        .Step_20   // Remove Lift comand
        .Step_03   // Rack Unlock Valve
        .Step_21   // Remove Unlock Comand
        .Step_04   // Lapbars Opening Valve -Y31008I
        .Step_22   // Lift comand
   RESTRAINTS_Left_Press_Switch_Series : BOOL := 1;
   RESTRAINTS_MainValve_PressTest : Valve_2_pos_monostable := (FeedBack_Type := 1, Discrepancy_Time := 2000, I_FeedBack_Data := 1, I_FeedBack_Status := 1, I_Output_Status := 1);
   RESTRAINTS_No_Alarms : BOOL := 1;
   RESTRAINTS_Open_Cycle_Ok : BOOL := 1;
   RESTRAINTS_Open_Postion : BOOL[64];
        [10]   // -B53201J
        [11]   // -B55001J
        [12]   // -B55007J
        [13]   // -B55101J
        [14]   // -B55107J
        [15]   // -B55201J
        [16]   // -B57001J
        [17]   // -B57007J
        [18]   // -B57101J
        [19]   // -B57107J
        [20]   // -B57201J
        [21]   // -B59001J
        [22]   // -B59007J
        [23]   // -B59101J
        [24]   // -B59107J
        [25]   // -B59201J
        [26]   // -B61001J
        [27]   // -B61007J
        [1]   // -B51001J
        [28]   // -B61101J
        [2]   // -B51007J
        [3]   // -B51101J
        [4]   // -B51107J
        [5]   // -B51201J
        [6]   // -B53001J
        [7]   // -B53007J
        [30]   // -B61201J
        [31]   // -B63001J
        [32]   // -B63007J
        [33]   // -B63101J
        [34]   // -B63107J
        [35]   // -B63201J
        [36]   // -B65001J
        [37]   // -B65007J
        [38]   // -B65101J
        [39]   // -B65007J
        [8]   // B53101J
        [9]   // B53107J
        [40]   // -B65201J
        [29]   // -B611017J
   RESTRAINTS_OpenComand : BOOL;   // Steps 01, 02, 03, 04
   RESTRAINTS_Opening : BOOL;
   Restraints_Permissive : Permissive := (All_Permissive_Ok := 1, BitsConditions := -1);
   Restraints_Permissive_Ok : BOOL := 1;
   Restraints_PermissiveLost : DINT := -2097153;
   RESTRAINTS_PressureSwitch_Working : BOOL := 1;
   RESTRAINTS_Rack : LapBar_Racks[41] := ([1].Input_Left.Discrepancy_Time := 3000, [1].Input_Left.Channel_A := 1, [1].Input_Left.Channel_B := 1, [1].Input_Left.Channel_A_Status := 1, [1].Input_Left.Channel_B_Status := 1, [1].Input_Left.O1 := 1, [1].Input_Right.Discrepancy_Time := 3000, [1].Input_Right.Channel_A := 1, [1].Input_Right.Channel_B := 1, [1].Input_Right.Channel_A_Status := 1, [1].Input_Right.Channel_B_Status := 1, [1].Input_Right.O1 := 1, [1].ON_Delay_Left.PRE := 500, [1].ON_Delay_Right.PRE := 500, [1].Memory_Left := 1, [1].Memory_Right := 1, [1].Memory_Left_Unlocked := 1, [1].Memory_Right_Unlocked := 1, [2].Input_Left.Discrepancy_Time := 3000, [2].Input_Left.Channel_A := 1, [2].Input_Left.Channel_B := 1, [2].Input_Left.Channel_A_Status := 1, [2].Input_Left.Channel_B_Status := 1, [2].Input_Left.O1 := 1, [2].Input_Right.Discrepancy_Time := 3000, [2].Input_Right.Channel_A := 1, [2].Input_Right.Channel_B := 1, [2].Input_Right.Channel_A_Status := 1, [2].Input_Right.Channel_B_Status := 1, [2].Input_Right.O1 := 1, [2].ON_Delay_Left.PRE := 500, [2].ON_Delay_Right.PRE := 500, [2].Memory_Left := 1, [2].Memory_Right := 1, [2].Memory_Left_Unlocked := 1, [2].Memory_Right_Unlocked := 1, [3].Input_Left.Discrepancy_Time := 3000, [3].Input_Left.Channel_A := 1, [3].Input_Left.Channel_B := 1, [3].Input_Left.Channel_A_Status := 1, [3].Input_Left.Channel_B_Status := 1, [3].Input_Left.O1 := 1, [3].Input_Right.Discrepancy_Time := 3000, [3].Input_Right.Channel_A := 1, [3].Input_Right.Channel_B := 1, [3].Input_Right.Channel_A_Status := 1, [3].Input_Right.Channel_B_Status := 1, [3].Input_Right.O1 := 1, [3].ON_Delay_Left.PRE := 500, [3].ON_Delay_Right.PRE := 500, [3].Memory_Left := 1, [3].Memory_Right := 1, [3].Memory_Left_Unlocked := 1, [3].Memory_Right_Unlocked := 1, [4].Input_Left.Discrepancy_Time := 3000, [4].Input_Left.Channel_A := 1, [4].Input_Left.Channel_B := 1, [4].Input_Left.Channel_A_Status := 1, [4].Input_Left.Channel_B_Status := 1, [4].Input_Left.O1 := 1,
        [4].Input_Right.Discrepancy_Time := 3000, [4].Input_Right.Channel_A := 1, [4].Input_Right.Channel_B := 1, [4].Input_Right.Channel_A_Status := 1, [4].Input_Right.Channel_B_Status := 1, [4].Input_Right.O1 := 1, [4].ON_Delay_Left.PRE := 500, [4].ON_Delay_Right.PRE := 500, [4].Memory_Left := 1, [4].Memory_Right := 1, [4].Memory_Left_Unlocked := 1, [4].Memory_Right_Unlocked := 1, [5].Input_Left.Discrepancy_Time := 3000, [5].Input_Left.Channel_A := 1, [5].Input_Left.Channel_B := 1, [5].Input_Left.Channel_A_Status := 1, [5].Input_Left.Channel_B_Status := 1, [5].Input_Left.O1 := 1, [5].Input_Right.Discrepancy_Time := 3000, [5].Input_Right.Channel_A := 1, [5].Input_Right.Channel_B := 1, [5].Input_Right.Channel_A_Status := 1, [5].Input_Right.Channel_B_Status := 1, [5].Input_Right.O1 := 1, [5].ON_Delay_Left.PRE := 500, [5].ON_Delay_Right.PRE := 500, [5].Memory_Left := 1, [5].Memory_Right := 1, [5].Memory_Left_Unlocked := 1, [5].Memory_Right_Unlocked := 1, [6].Input_Left.Discrepancy_Time := 3000, [6].Input_Left.Channel_A := 1, [6].Input_Left.Channel_B := 1, [6].Input_Left.Channel_A_Status := 1, [6].Input_Left.Channel_B_Status := 1, [6].Input_Left.O1 := 1, [6].Input_Right.Discrepancy_Time := 3000, [6].Input_Right.Channel_A := 1, [6].Input_Right.Channel_B := 1, [6].Input_Right.Channel_A_Status := 1, [6].Input_Right.Channel_B_Status := 1, [6].Input_Right.O1 := 1, [6].ON_Delay_Left.PRE := 500, [6].ON_Delay_Right.PRE := 500, [6].Memory_Left := 1, [6].Memory_Right := 1, [6].Memory_Left_Unlocked := 1, [6].Memory_Right_Unlocked := 1, [7].Input_Left.Discrepancy_Time := 3000, [7].Input_Left.Channel_A := 1, [7].Input_Left.Channel_B := 1, [7].Input_Left.Channel_A_Status := 1, [7].Input_Left.Channel_B_Status := 1, [7].Input_Left.O1 := 1, [7].Input_Right.Discrepancy_Time := 3000, [7].Input_Right.Channel_A := 1, [7].Input_Right.Channel_B := 1, [7].Input_Right.Channel_A_Status := 1, [7].Input_Right.Channel_B_Status := 1, [7].Input_Right.O1 := 1,
        [7].ON_Delay_Left.PRE := 500, [7].ON_Delay_Right.PRE := 500, [7].Memory_Left := 1, [7].Memory_Right := 1, [7].Memory_Left_Unlocked := 1, [7].Memory_Right_Unlocked := 1, [8].Input_Left.Discrepancy_Time := 3000, [8].Input_Left.Channel_A := 1, [8].Input_Left.Channel_B := 1, [8].Input_Left.Channel_A_Status := 1, [8].Input_Left.Channel_B_Status := 1, [8].Input_Left.O1 := 1, [8].Input_Right.Discrepancy_Time := 3000, [8].Input_Right.Channel_A := 1, [8].Input_Right.Channel_B := 1, [8].Input_Right.Channel_A_Status := 1, [8].Input_Right.Channel_B_Status := 1, [8].Input_Right.O1 := 1, [8].ON_Delay_Left.PRE := 500, [8].ON_Delay_Right.PRE := 500, [8].Memory_Left := 1, [8].Memory_Right := 1, [8].Memory_Left_Unlocked := 1, [8].Memory_Right_Unlocked := 1, [9].Input_Left.Discrepancy_Time := 3000, [9].Input_Left.Channel_A := 1, [9].Input_Left.Channel_B := 1, [9].Input_Left.Channel_A_Status := 1, [9].Input_Left.Channel_B_Status := 1, [9].Input_Left.O1 := 1, [9].Input_Right.Discrepancy_Time := 3000, [9].Input_Right.Channel_A_Status := 1, [9].Input_Right.Channel_B_Status := 1, [9].ON_Delay_Left.PRE := 500, [9].ON_Delay_Right.PRE := 500, [9].Memory_Left := 1, [9].Memory_Right := 1, [9].Memory_Left_Unlocked := 1, [9].Memory_Right_Unlocked := 1, [10].Input_Left.Discrepancy_Time := 3000, [10].Input_Left.Channel_A := 1, [10].Input_Left.Channel_B := 1, [10].Input_Left.Channel_A_Status := 1, [10].Input_Left.Channel_B_Status := 1, [10].Input_Left.O1 := 1, [10].Input_Right.Discrepancy_Time := 3000, [10].Input_Right.Channel_A := 1, [10].Input_Right.Channel_B := 1, [10].Input_Right.Channel_A_Status := 1, [10].Input_Right.Channel_B_Status := 1, [10].Input_Right.O1 := 1, [10].ON_Delay_Left.PRE := 500, [10].ON_Delay_Right.PRE := 500, [10].Memory_Left := 1, [10].Memory_Right := 1, [10].Memory_Left_Unlocked := 1, [10].Memory_Right_Unlocked := 1, [11].Input_Left.Discrepancy_Time := 3000, [11].Input_Left.Channel_A := 1, [11].Input_Left.Channel_B := 1,
        [11].Input_Left.Channel_A_Status := 1, [11].Input_Left.Channel_B_Status := 1, [11].Input_Left.O1 := 1, [11].Input_Right.Discrepancy_Time := 3000, [11].Input_Right.Channel_A := 1, [11].Input_Right.Channel_B := 1, [11].Input_Right.Channel_A_Status := 1, [11].Input_Right.Channel_B_Status := 1, [11].Input_Right.O1 := 1, [11].ON_Delay_Left.PRE := 500, [11].ON_Delay_Right.PRE := 500, [11].Memory_Left := 1, [11].Memory_Right := 1, [11].Memory_Left_Unlocked := 1, [11].Memory_Right_Unlocked := 1, [12].Input_Left.Discrepancy_Time := 3000, [12].Input_Left.Channel_A := 1, [12].Input_Left.Channel_B := 1, [12].Input_Left.Channel_A_Status := 1, [12].Input_Left.Channel_B_Status := 1, [12].Input_Left.O1 := 1, [12].Input_Right.Discrepancy_Time := 3000, [12].Input_Right.Channel_A := 1, [12].Input_Right.Channel_B := 1, [12].Input_Right.Channel_A_Status := 1, [12].Input_Right.Channel_B_Status := 1, [12].Input_Right.O1 := 1, [12].ON_Delay_Left.PRE := 500, [12].ON_Delay_Right.PRE := 500, [12].Memory_Left := 1, [12].Memory_Right := 1, [12].Memory_Left_Unlocked := 1, [12].Memory_Right_Unlocked := 1, [13].Input_Left.Discrepancy_Time := 3000, [13].Input_Left.Channel_A := 1, [13].Input_Left.Channel_B := 1, [13].Input_Left.Channel_A_Status := 1, [13].Input_Left.Channel_B_Status := 1, [13].Input_Left.O1 := 1, [13].Input_Right.Discrepancy_Time := 3000, [13].Input_Right.Channel_A := 1, [13].Input_Right.Channel_B := 1, [13].Input_Right.Channel_A_Status := 1, [13].Input_Right.Channel_B_Status := 1, [13].Input_Right.O1 := 1, [13].ON_Delay_Left.PRE := 500, [13].ON_Delay_Right.PRE := 500, [13].Memory_Left := 1, [13].Memory_Right := 1, [13].Memory_Left_Unlocked := 1, [13].Memory_Right_Unlocked := 1, [14].Input_Left.Discrepancy_Time := 3000, [14].Input_Left.Channel_A := 1, [14].Input_Left.Channel_B := 1, [14].Input_Left.Channel_A_Status := 1, [14].Input_Left.Channel_B_Status := 1, [14].Input_Left.O1 := 1, [14].Input_Right.Discrepancy_Time := 3000, [14].Input_Right.Channel_A := 1, [14].Input_Right.Channel_B := 1,
        [14].Input_Right.Channel_A_Status := 1, [14].Input_Right.Channel_B_Status := 1, [14].Input_Right.O1 := 1, [14].ON_Delay_Left.PRE := 500, [14].ON_Delay_Right.PRE := 500, [14].Memory_Left := 1, [14].Memory_Right := 1, [14].Memory_Left_Unlocked := 1, [14].Memory_Right_Unlocked := 1, [15].Input_Left.Discrepancy_Time := 3000, [15].Input_Left.Channel_A := 1, [15].Input_Left.Channel_B := 1, [15].Input_Left.Channel_A_Status := 1, [15].Input_Left.Channel_B_Status := 1, [15].Input_Left.O1 := 1, [15].Input_Right.Discrepancy_Time := 3000, [15].Input_Right.Channel_A := 1, [15].Input_Right.Channel_B := 1, [15].Input_Right.Channel_A_Status := 1, [15].Input_Right.Channel_B_Status := 1, [15].Input_Right.O1 := 1, [15].ON_Delay_Left.PRE := 500, [15].ON_Delay_Right.PRE := 500, [15].Memory_Left := 1, [15].Memory_Right := 1, [15].Memory_Left_Unlocked := 1, [15].Memory_Right_Unlocked := 1, [16].Input_Left.Discrepancy_Time := 3000, [16].Input_Left.Channel_A := 1, [16].Input_Left.Channel_B := 1, [16].Input_Left.Channel_A_Status := 1, [16].Input_Left.Channel_B_Status := 1, [16].Input_Left.O1 := 1, [16].Input_Right.Discrepancy_Time := 3000, [16].Input_Right.Channel_A := 1, [16].Input_Right.Channel_B := 1, [16].Input_Right.Channel_A_Status := 1, [16].Input_Right.Channel_B_Status := 1, [16].Input_Right.O1 := 1, [16].ON_Delay_Left.PRE := 500, [16].ON_Delay_Right.PRE := 500, [16].Memory_Left := 1, [16].Memory_Right := 1, [16].Memory_Left_Unlocked := 1, [16].Memory_Right_Unlocked := 1, [17].Input_Left.Discrepancy_Time := 3000, [17].Input_Left.Channel_A := 1, [17].Input_Left.Channel_B := 1, [17].Input_Left.Channel_A_Status := 1, [17].Input_Left.Channel_B_Status := 1, [17].Input_Left.O1 := 1, [17].Input_Right.Discrepancy_Time := 3000, [17].Input_Right.Channel_A := 1, [17].Input_Right.Channel_B := 1, [17].Input_Right.Channel_A_Status := 1, [17].Input_Right.Channel_B_Status := 1, [17].Input_Right.O1 := 1, [17].ON_Delay_Left.PRE := 500, [17].ON_Delay_Right.PRE := 500, [17].Memory_Left := 1,
        [17].Memory_Right := 1, [18].Input_Left.Discrepancy_Time := 3000, [18].Input_Left.Channel_A := 1, [18].Input_Left.Channel_B := 1, [18].Input_Left.Channel_A_Status := 1, [18].Input_Left.Channel_B_Status := 1, [18].Input_Left.O1 := 1, [18].Input_Right.Discrepancy_Time := 3000, [18].Input_Right.Channel_A := 1, [18].Input_Right.Channel_B := 1, [18].Input_Right.Channel_A_Status := 1, [18].Input_Right.Channel_B_Status := 1, [18].Input_Right.O1 := 1, [18].ON_Delay_Left.PRE := 500, [18].ON_Delay_Right.PRE := 500, [18].Memory_Left := 1, [18].Memory_Right := 1, [19].Input_Left.Discrepancy_Time := 3000, [19].Input_Left.Channel_A := 1, [19].Input_Left.Channel_B := 1, [19].Input_Left.Channel_A_Status := 1, [19].Input_Left.Channel_B_Status := 1, [19].Input_Left.O1 := 1, [19].Input_Right.Discrepancy_Time := 3000, [19].Input_Right.Channel_A := 1, [19].Input_Right.Channel_B := 1, [19].Input_Right.Channel_A_Status := 1, [19].Input_Right.Channel_B_Status := 1, [19].Input_Right.O1 := 1, [19].ON_Delay_Left.PRE := 500, [19].ON_Delay_Right.PRE := 500, [19].Memory_Left := 1, [19].Memory_Right := 1, [20].Input_Left.Discrepancy_Time := 3000, [20].Input_Left.Channel_A := 1, [20].Input_Left.Channel_B := 1, [20].Input_Left.Channel_A_Status := 1, [20].Input_Left.Channel_B_Status := 1, [20].Input_Left.O1 := 1, [20].Input_Right.Discrepancy_Time := 3000, [20].Input_Right.Channel_A := 1, [20].Input_Right.Channel_B := 1, [20].Input_Right.Channel_A_Status := 1, [20].Input_Right.Channel_B_Status := 1, [20].Input_Right.O1 := 1, [20].ON_Delay_Left.PRE := 500, [20].ON_Delay_Right.PRE := 500, [20].Memory_Left := 1, [20].Memory_Right := 1, [21].Input_Left.Discrepancy_Time := 3000, [21].Input_Left.Channel_A := 1, [21].Input_Left.Channel_B := 1, [21].Input_Left.Channel_A_Status := 1, [21].Input_Left.Channel_B_Status := 1, [21].Input_Left.O1 := 1, [21].Input_Right.Discrepancy_Time := 3000, [21].Input_Right.Channel_A := 1, [21].Input_Right.Channel_B := 1, [21].Input_Right.Channel_A_Status := 1, [21].Input_Right.Channel_B_Status := 1,
        [21].Input_Right.O1 := 1, [21].ON_Delay_Left.PRE := 500, [21].ON_Delay_Right.PRE := 500, [21].Memory_Left := 1, [21].Memory_Right := 1, [22].Input_Left.Discrepancy_Time := 3000, [22].Input_Left.Channel_A := 1, [22].Input_Left.Channel_B := 1, [22].Input_Left.Channel_A_Status := 1, [22].Input_Left.Channel_B_Status := 1, [22].Input_Left.O1 := 1, [22].Input_Right.Discrepancy_Time := 3000, [22].Input_Right.Channel_A := 1, [22].Input_Right.Channel_B := 1, [22].Input_Right.Channel_A_Status := 1, [22].Input_Right.Channel_B_Status := 1, [22].Input_Right.O1 := 1, [22].ON_Delay_Left.PRE := 500, [22].ON_Delay_Right.PRE := 500, [22].Memory_Left := 1, [22].Memory_Right := 1, [23].Input_Left.Discrepancy_Time := 3000, [23].Input_Left.Channel_A := 1, [23].Input_Left.Channel_B := 1, [23].Input_Left.Channel_A_Status := 1, [23].Input_Left.Channel_B_Status := 1, [23].Input_Left.O1 := 1, [23].Input_Right.Discrepancy_Time := 3000, [23].Input_Right.Channel_A := 1, [23].Input_Right.Channel_B := 1, [23].Input_Right.Channel_A_Status := 1, [23].Input_Right.Channel_B_Status := 1, [23].Input_Right.O1 := 1, [23].ON_Delay_Left.PRE := 500, [23].ON_Delay_Right.PRE := 500, [23].Memory_Left := 1, [23].Memory_Right := 1, [24].Input_Left.Discrepancy_Time := 3000, [24].Input_Left.Channel_A := 1, [24].Input_Left.Channel_B := 1, [24].Input_Left.Channel_A_Status := 1, [24].Input_Left.Channel_B_Status := 1, [24].Input_Left.O1 := 1, [24].Input_Right.Discrepancy_Time := 3000, [24].Input_Right.Channel_A := 1, [24].Input_Right.Channel_B := 1, [24].Input_Right.Channel_A_Status := 1, [24].Input_Right.Channel_B_Status := 1, [24].Input_Right.O1 := 1, [24].ON_Delay_Left.PRE := 500, [24].ON_Delay_Right.PRE := 500, [24].Memory_Left := 1, [24].Memory_Right := 1, [25].Input_Left.Discrepancy_Time := 3000, [25].Input_Left.Channel_A := 1, [25].Input_Left.Channel_B := 1, [25].Input_Left.Channel_A_Status := 1, [25].Input_Left.Channel_B_Status := 1, [25].Input_Left.O1 := 1, [25].Input_Right.Discrepancy_Time := 3000,
        [25].Input_Right.Channel_A := 1, [25].Input_Right.Channel_B := 1, [25].Input_Right.Channel_A_Status := 1, [25].Input_Right.Channel_B_Status := 1, [25].Input_Right.O1 := 1, [25].ON_Delay_Left.PRE := 500, [25].ON_Delay_Right.PRE := 500, [25].Memory_Left := 1, [25].Memory_Right := 1, [26].Input_Left.Discrepancy_Time := 3000, [26].Input_Left.Channel_A := 1, [26].Input_Left.Channel_B := 1, [26].Input_Left.Channel_A_Status := 1, [26].Input_Left.Channel_B_Status := 1, [26].Input_Left.O1 := 1, [26].Input_Right.Discrepancy_Time := 3000, [26].Input_Right.Channel_A := 1, [26].Input_Right.Channel_B := 1, [26].Input_Right.Channel_A_Status := 1, [26].Input_Right.Channel_B_Status := 1, [26].Input_Right.O1 := 1, [26].ON_Delay_Left.PRE := 500, [26].ON_Delay_Right.PRE := 500, [26].Memory_Left := 1, [26].Memory_Right := 1, [27].Input_Left.Discrepancy_Time := 3000, [27].Input_Left.Channel_A := 1, [27].Input_Left.Channel_B := 1, [27].Input_Left.Channel_A_Status := 1, [27].Input_Left.Channel_B_Status := 1, [27].Input_Left.O1 := 1, [27].Input_Right.Discrepancy_Time := 3000, [27].Input_Right.Channel_A := 1, [27].Input_Right.Channel_B := 1, [27].Input_Right.Channel_A_Status := 1, [27].Input_Right.Channel_B_Status := 1, [27].Input_Right.O1 := 1, [27].ON_Delay_Left.PRE := 500, [27].ON_Delay_Right.PRE := 500, [27].Memory_Left := 1, [27].Memory_Right := 1, [28].Input_Left.Discrepancy_Time := 3000, [28].Input_Left.Channel_A := 1, [28].Input_Left.Channel_B := 1, [28].Input_Left.Channel_A_Status := 1, [28].Input_Left.Channel_B_Status := 1, [28].Input_Left.O1 := 1, [28].Input_Right.Discrepancy_Time := 3000, [28].Input_Right.Channel_A := 1, [28].Input_Right.Channel_B := 1, [28].Input_Right.Channel_A_Status := 1, [28].Input_Right.Channel_B_Status := 1, [28].Input_Right.O1 := 1, [28].ON_Delay_Left.PRE := 500, [28].ON_Delay_Right.PRE := 500, [28].Memory_Left := 1, [28].Memory_Right := 1, [29].Input_Left.Discrepancy_Time := 3000, [29].Input_Left.Channel_A := 1, [29].Input_Left.Channel_B := 1,
        [29].Input_Left.Channel_A_Status := 1, [29].Input_Left.Channel_B_Status := 1, [29].Input_Left.O1 := 1, [29].Input_Right.Discrepancy_Time := 3000, [29].Input_Right.Channel_A := 1, [29].Input_Right.Channel_B := 1, [29].Input_Right.Channel_A_Status := 1, [29].Input_Right.Channel_B_Status := 1, [29].Input_Right.O1 := 1, [29].ON_Delay_Left.PRE := 500, [29].ON_Delay_Right.PRE := 500, [29].Memory_Left := 1, [29].Memory_Right := 1, [30].Input_Left.Discrepancy_Time := 3000, [30].Input_Left.Channel_A := 1, [30].Input_Left.Channel_B := 1, [30].Input_Left.Channel_A_Status := 1, [30].Input_Left.Channel_B_Status := 1, [30].Input_Left.O1 := 1, [30].Input_Right.Discrepancy_Time := 3000, [30].Input_Right.Channel_A := 1, [30].Input_Right.Channel_B := 1, [30].Input_Right.Channel_A_Status := 1, [30].Input_Right.Channel_B_Status := 1, [30].Input_Right.O1 := 1, [30].ON_Delay_Left.PRE := 500, [30].ON_Delay_Right.PRE := 500, [30].Memory_Left := 1, [30].Memory_Right := 1, [31].Input_Left.Discrepancy_Time := 3000, [31].Input_Left.Channel_A := 1, [31].Input_Left.Channel_B := 1, [31].Input_Left.Channel_A_Status := 1, [31].Input_Left.Channel_B_Status := 1, [31].Input_Left.O1 := 1, [31].Input_Right.Discrepancy_Time := 3000, [31].Input_Right.Channel_A := 1, [31].Input_Right.Channel_B := 1, [31].Input_Right.Channel_A_Status := 1, [31].Input_Right.Channel_B_Status := 1, [31].Input_Right.O1 := 1, [31].ON_Delay_Left.PRE := 500, [31].ON_Delay_Right.PRE := 500, [31].Memory_Left := 1, [31].Memory_Right := 1, [32].Input_Left.Discrepancy_Time := 3000, [32].Input_Left.Channel_A := 1, [32].Input_Left.Channel_B := 1, [32].Input_Left.Channel_A_Status := 1, [32].Input_Left.Channel_B_Status := 1, [32].Input_Left.O1 := 1, [32].Input_Right.Discrepancy_Time := 3000, [32].Input_Right.Channel_A := 1, [32].Input_Right.Channel_B := 1, [32].Input_Right.Channel_A_Status := 1, [32].Input_Right.Channel_B_Status := 1, [32].Input_Right.O1 := 1, [32].ON_Delay_Left.PRE := 500, [32].ON_Delay_Right.PRE := 500, [32].Memory_Left := 1,
        [32].Memory_Right := 1, [33].Input_Left.Discrepancy_Time := 3000, [33].Input_Left.Channel_A := 1, [33].Input_Left.Channel_B := 1, [33].Input_Left.Channel_A_Status := 1, [33].Input_Left.Channel_B_Status := 1, [33].Input_Left.O1 := 1, [33].Input_Right.Discrepancy_Time := 3000, [33].Input_Right.Channel_A := 1, [33].Input_Right.Channel_B := 1, [33].Input_Right.Channel_A_Status := 1, [33].Input_Right.Channel_B_Status := 1, [33].Input_Right.O1 := 1, [33].ON_Delay_Left.PRE := 500, [33].ON_Delay_Right.PRE := 500, [33].Memory_Left := 1, [33].Memory_Right := 1, [34].Input_Left.Discrepancy_Time := 3000, [34].Input_Left.Channel_A := 1, [34].Input_Left.Channel_B := 1, [34].Input_Left.Channel_A_Status := 1, [34].Input_Left.Channel_B_Status := 1, [34].Input_Left.O1 := 1, [34].Input_Right.Discrepancy_Time := 3000, [34].Input_Right.Channel_A := 1, [34].Input_Right.Channel_B := 1, [34].Input_Right.Channel_A_Status := 1, [34].Input_Right.Channel_B_Status := 1, [34].Input_Right.O1 := 1, [34].ON_Delay_Left.PRE := 500, [34].ON_Delay_Right.PRE := 500, [34].Memory_Left := 1, [34].Memory_Right := 1, [35].Input_Left.Discrepancy_Time := 3000, [35].Input_Left.Channel_A := 1, [35].Input_Left.Channel_B := 1, [35].Input_Left.Channel_A_Status := 1, [35].Input_Left.Channel_B_Status := 1, [35].Input_Left.O1 := 1, [35].Input_Right.Discrepancy_Time := 3000, [35].Input_Right.Channel_A := 1, [35].Input_Right.Channel_B := 1, [35].Input_Right.Channel_A_Status := 1, [35].Input_Right.Channel_B_Status := 1, [35].Input_Right.O1 := 1, [35].ON_Delay_Left.PRE := 500, [35].ON_Delay_Right.PRE := 500, [35].Memory_Left := 1, [35].Memory_Right := 1, [36].Input_Left.Discrepancy_Time := 3000, [36].Input_Left.Channel_A := 1, [36].Input_Left.Channel_B := 1, [36].Input_Left.Channel_A_Status := 1, [36].Input_Left.Channel_B_Status := 1, [36].Input_Left.O1 := 1, [36].Input_Right.Discrepancy_Time := 3000, [36].Input_Right.Channel_A := 1, [36].Input_Right.Channel_B := 1, [36].Input_Right.Channel_A_Status := 1, [36].Input_Right.Channel_B_Status := 1,
        [36].Input_Right.O1 := 1, [36].ON_Delay_Left.PRE := 500, [36].ON_Delay_Right.PRE := 500, [36].Memory_Left := 1, [36].Memory_Right := 1, [37].Input_Left.Discrepancy_Time := 3000, [37].Input_Left.Channel_A := 1, [37].Input_Left.Channel_B := 1, [37].Input_Left.Channel_A_Status := 1, [37].Input_Left.Channel_B_Status := 1, [37].Input_Left.O1 := 1, [37].Input_Right.Discrepancy_Time := 3000, [37].Input_Right.Channel_A := 1, [37].Input_Right.Channel_B := 1, [37].Input_Right.Channel_A_Status := 1, [37].Input_Right.Channel_B_Status := 1, [37].Input_Right.O1 := 1, [37].ON_Delay_Left.PRE := 500, [37].ON_Delay_Right.PRE := 500, [37].Memory_Left := 1, [37].Memory_Right := 1, [38].Input_Left.Discrepancy_Time := 3000, [38].Input_Left.Channel_A := 1, [38].Input_Left.Channel_B := 1, [38].Input_Left.Channel_A_Status := 1, [38].Input_Left.Channel_B_Status := 1, [38].Input_Left.O1 := 1, [38].Input_Right.Discrepancy_Time := 3000, [38].Input_Right.Channel_A := 1, [38].Input_Right.Channel_B := 1, [38].Input_Right.Channel_A_Status := 1, [38].Input_Right.Channel_B_Status := 1, [38].Input_Right.O1 := 1, [38].ON_Delay_Left.PRE := 500, [38].ON_Delay_Right.PRE := 500, [38].Memory_Left := 1, [38].Memory_Right := 1, [39].Input_Left.Discrepancy_Time := 3000, [39].Input_Left.Channel_A := 1, [39].Input_Left.Channel_B := 1, [39].Input_Left.Channel_A_Status := 1, [39].Input_Left.Channel_B_Status := 1, [39].Input_Left.O1 := 1, [39].Input_Right.Discrepancy_Time := 3000, [39].Input_Right.Channel_A := 1, [39].Input_Right.Channel_B := 1, [39].Input_Right.Channel_A_Status := 1, [39].Input_Right.Channel_B_Status := 1, [39].Input_Right.O1 := 1, [39].ON_Delay_Left.PRE := 500, [39].ON_Delay_Right.PRE := 500, [39].Memory_Left := 1, [39].Memory_Right := 1, [40].Input_Left.Discrepancy_Time := 3000, [40].Input_Left.Channel_A := 1, [40].Input_Left.Channel_B := 1, [40].Input_Left.Channel_A_Status := 1, [40].Input_Left.Channel_B_Status := 1, [40].Input_Left.O1 := 1, [40].Input_Right.Discrepancy_Time := 3000,
        [40].Input_Right.Channel_A := 1, [40].Input_Right.Channel_B := 1, [40].Input_Right.Channel_A_Status := 1, [40].Input_Right.Channel_B_Status := 1, [40].Input_Right.O1 := 1, [40].ON_Delay_Left.PRE := 500, [40].ON_Delay_Right.PRE := 500, [40].Memory_Left := 1, [40].Memory_Right := 1);
        [10].Input_Left   // -A53702I
        [1].Input_Left   // -A51302I
        [10].Input_Right   // -A53707I
        [1].Input_Right   // -A51307I
        [2].Input_Left   // -A51402I
        [11].Input_Left   // -A55302I
        [2].Input_Right   // -A51407I
        [11].Input_Right   // -A55307I
        [12].Input_Left   // -A55402I
        [12].Input_Right   // -A55407I
        [13].Input_Left   // -A55502I
        [3].Input_Left   // -A51502I
        [13].Input_Right   // -A55507I
        [3].Input_Right   // -A51507I
        [4].Input_Left   // -A51602I
        [4].Input_Right   // -A51607I
        [5].Input_Left   // -A51702I
        [5].Input_Right   // -A51707I
        [6].Input_Left   // -A53302I
        [6].Input_Right   // -A53307I
        [7].Input_Left   // -A53402I
        [14].Input_Left   // -A55602I
        [7].Input_Right   // -A534027I
        [14].Input_Right   // -A55607I
        [15].Input_Left   // -A55702I
        [15].Input_Right   // -A55707I
        [8].Input_Left   // -A53502I
        [8].Input_Right   // -A53507I
        [9].Input_Left   // -A53602I
        [9].Input_Right   // -A53607I
        [16].Input_Left   // -A57402I
        [16].Input_Right   // -A57407I
        [17].Input_Left   // -A57402I
        [17].Input_Right   // -A57407I
        [18].Input_Left   // -A57502I
        [18].Input_Right   // -A57507I
        [19].Input_Left   // -A57602I
        [19].Input_Right   // -A57607I
        [20].Input_Left   // -A57702I
        [20].Input_Right   // -A57707I
        [21].Input_Left   // -A59302I
        [21].Input_Right   // -A59307I
        [22].Input_Left   // -A59402I
        [22].Input_Right   // -A59407I
        [23].Input_Left   // -A59502I
        [23].Input_Right   // -A59507I
        [24].Input_Left   // -A59602I
        [24].Input_Right   // -A59607I
        [25].Input_Left   // -A59702I
        [25].Input_Right   // -A59707I
        [26].Input_Left   // -A61302I
        [26].Input_Right   // -A61307I
        [27].Input_Left   // -A61402I
        [27].Input_Right   // -A61407I
        [28].Input_Left   // -A61502I
        [28].Input_Right   // -A61507I
        [29].Input_Left   // -A61602I
        [29].Input_Right   // -A61607I
        [30].Input_Left   // -A61702I
        [30].Input_Right   // -A61707I
        [31].Input_Left   // -A63302I
        [31].Input_Right   // -A63307I
        [32].Input_Left   // -A63402I
        [32].Input_Right   // -A63402I
        [33].Input_Left   // -A63502I
        [33].Input_Right   // -A63507I
        [34].Input_Left   // -A63602I
        [34].Input_Right   // -A63607I
        [35].Input_Left   // -A63702I
        [35].Input_Right   // -A63707I
        [36].Input_Left   // -A65302I
        [36].Input_Right   // -A65307I
        [37].Input_Left   // -A65402I
        [37].Input_Right   // -A65407I
        [38].Input_Left   // -A65502I
        [38].Input_Right   // -A65507I
        [39].Input_Left   // -A65602I
        [39].Input_Right   // -A65607I
        [40].Input_Left   // -A65702I
        [40].Input_Right   // -A65707I
   RESTRAINTS_Rack_Sector : BOOL;
   RESTRAINTS_Rack_Sector_A_ON : BOOL := 1;
   RESTRAINTS_Rack_Sector_ON : BOOL := 1;
   RESTRAINTS_Right_Press_Switch_Series : BOOL := 1;
   RESTRAINTS_Sector : LapBars_Sector[9] := ([1].Sensors_ChA := 1, [1].Sensors_ChB := 1, [1].LapBar_Open_Close := 1, [1].Input_Status := 1, [1].Sensor_ChA_Open_Memory := 1, [1].Sensor_ChB_Open_Memory := 1, [1].I_LB_PressureSwitch_Valve_Right_Open := 1, [1].I_LB_PressureSwitch_Valve_Left_Open := 1, [1].All_Rack_Memory_Signal_ON := 1, [1].RESTRAINTS_Rack_Sector_ON := 1, [1].I_Close_Position.ChannelA := 1, [1].I_Close_Position.ChannelB := 1, [1].I_Close_Position.InputStatus := 1, [1].I_Close_Position.SafetyFunction := 41, [1].I_Close_Position.DiscrepancyTime := 3000, [1].I_Close_Position.O1 := 1, [1].I_Close_Position.IS := 1, [1].I_Sector_Disable_Switch.Dual_Chanel_Monitor.ChannelB := 1, [1].I_Sector_Disable_Switch.Dual_Chanel_Monitor.InputStatus := 1, [1].I_Sector_Disable_Switch.Dual_Chanel_Monitor.SafetyFunction := 41, [1].I_Sector_Disable_Switch.Dual_Chanel_Monitor.InputType := 2, [1].I_Sector_Disable_Switch.Dual_Chanel_Monitor.DiscrepancyTime := 3000, [1].I_Sector_Disable_Switch.Dual_Chanel_Monitor.IS := 1, [1].I_Sector_Disable_Switch.Status := 1, [1].O_Unlock_Valve_Left.FeedBack_Type := 1, [1].O_Unlock_Valve_Left.Discrepancy_Time := 3000, [1].O_Unlock_Valve_Left.I_FeedBack_Data := 1, [1].O_Unlock_Valve_Left.I_FeedBack_Status := 1, [1].O_Unlock_Valve_Left.I_Output_Status := 1, [1].O_Unlock_Valve_Right.FeedBack_Type := 1, [1].O_Unlock_Valve_Right.Discrepancy_Time := 3000, [1].O_Unlock_Valve_Right.I_FeedBack_Data := 1, [1].O_Unlock_Valve_Right.I_FeedBack_Status := 1, [1].O_Unlock_Valve_Right.I_Output_Status := 1, [2].Sensors_ChA := 1, [2].Sensors_ChB := 1, [2].LapBar_Open_Close := 1, [2].Input_Status := 1, [2].Sensor_ChA_Open_Memory := 1, [2].Sensor_ChB_Open_Memory := 1, [2].I_LB_PressureSwitch_Valve_Right_Open := 1, [2].I_LB_PressureSwitch_Valve_Left_Open := 1, [2].All_Rack_Memory_Signal_ON := 1, [2].RESTRAINTS_Rack_Sector_ON := 1, [2].I_Close_Position.ChannelA := 1, [2].I_Close_Position.ChannelB := 1, [2].I_Close_Position.InputStatus := 1, [2].I_Close_Position.SafetyFunction := 41, [2].I_Close_Position.DiscrepancyTime := 3000, [2].I_Close_Position.O1 := 1, [2].I_Close_Position.IS := 1, [2].I_Sector_Disable_Switch.Dual_Chanel_Monitor.ChannelB := 1, [2].I_Sector_Disable_Switch.Dual_Chanel_Monitor.InputStatus := 1, [2].I_Sector_Disable_Switch.Dual_Chanel_Monitor.SafetyFunction := 41, [2].I_Sector_Disable_Switch.Dual_Chanel_Monitor.InputType := 2, [2].I_Sector_Disable_Switch.Dual_Chanel_Monitor.DiscrepancyTime := 3000, [2].I_Sector_Disable_Switch.Dual_Chanel_Monitor.IS := 1, [2].I_Sector_Disable_Switch.Status := 1, [2].O_Unlock_Valve_Left.FeedBack_Type := 1, [2].O_Unlock_Valve_Left.Discrepancy_Time := 3000,
        [2].O_Unlock_Valve_Left.I_FeedBack_Data := 1, [2].O_Unlock_Valve_Left.I_FeedBack_Status := 1, [2].O_Unlock_Valve_Left.I_Output_Status := 1, [2].O_Unlock_Valve_Right.FeedBack_Type := 1, [2].O_Unlock_Valve_Right.Discrepancy_Time := 3000, [2].O_Unlock_Valve_Right.I_FeedBack_Data := 1, [2].O_Unlock_Valve_Right.I_FeedBack_Status := 1, [2].O_Unlock_Valve_Right.I_Output_Status := 1, [3].Sensors_ChA := 1, [3].Sensors_ChB := 1, [3].LapBar_Open_Close := 1, [3].Input_Status := 1, [3].Sensor_ChA_Open_Memory := 1, [3].Sensor_ChB_Open_Memory := 1, [3].I_LB_PressureSwitch_Valve_Right_Open := 1, [3].I_LB_PressureSwitch_Valve_Left_Open := 1, [3].All_Rack_Memory_Signal_ON := 1, [3].RESTRAINTS_Rack_Sector_ON := 1, [3].I_Close_Position.ChannelA := 1, [3].I_Close_Position.ChannelB := 1, [3].I_Close_Position.InputStatus := 1, [3].I_Close_Position.SafetyFunction := 41, [3].I_Close_Position.DiscrepancyTime := 3000, [3].I_Close_Position.O1 := 1, [3].I_Close_Position.IS := 1, [3].I_Sector_Disable_Switch.Dual_Chanel_Monitor.ChannelB := 1, [3].I_Sector_Disable_Switch.Dual_Chanel_Monitor.InputStatus := 1, [3].I_Sector_Disable_Switch.Dual_Chanel_Monitor.SafetyFunction := 41, [3].I_Sector_Disable_Switch.Dual_Chanel_Monitor.InputType := 2, [3].I_Sector_Disable_Switch.Dual_Chanel_Monitor.DiscrepancyTime := 3000, [3].I_Sector_Disable_Switch.Dual_Chanel_Monitor.IS := 1, [3].I_Sector_Disable_Switch.Status := 1, [3].O_Unlock_Valve_Left.FeedBack_Type := 1, [3].O_Unlock_Valve_Left.Discrepancy_Time := 3000, [3].O_Unlock_Valve_Left.I_FeedBack_Data := 1, [3].O_Unlock_Valve_Left.I_FeedBack_Status := 1, [3].O_Unlock_Valve_Left.I_Output_Status := 1, [3].O_Unlock_Valve_Right.FeedBack_Type := 1, [3].O_Unlock_Valve_Right.Discrepancy_Time := 3000, [3].O_Unlock_Valve_Right.I_FeedBack_Data := 1, [3].O_Unlock_Valve_Right.I_FeedBack_Status := 1, [3].O_Unlock_Valve_Right.I_Output_Status := 1, [4].Sensors_ChA := 1, [4].Sensors_ChB := 1, [4].LapBar_Open_Close := 1, [4].Input_Status := 1, [4].Sensor_ChA_Open_Memory := 1, [4].Sensor_ChB_Open_Memory := 1, [4].I_LB_PressureSwitch_Valve_Right_Open := 1, [4].I_LB_PressureSwitch_Valve_Left_Open := 1, [4].All_Rack_Memory_Signal_ON := 1, [4].RESTRAINTS_Rack_Sector_ON := 1, [4].I_Close_Position.ChannelA := 1, [4].I_Close_Position.ChannelB := 1, [4].I_Close_Position.InputStatus := 1, [4].I_Close_Position.SafetyFunction := 41, [4].I_Close_Position.DiscrepancyTime := 3000, [4].I_Close_Position.O1 := 1, [4].I_Close_Position.IS := 1, [4].I_Sector_Disable_Switch.Dual_Chanel_Monitor.ChannelB := 1,
        [4].I_Sector_Disable_Switch.Dual_Chanel_Monitor.InputStatus := 1, [4].I_Sector_Disable_Switch.Dual_Chanel_Monitor.SafetyFunction := 41, [4].I_Sector_Disable_Switch.Dual_Chanel_Monitor.InputType := 2, [4].I_Sector_Disable_Switch.Dual_Chanel_Monitor.DiscrepancyTime := 3000, [4].I_Sector_Disable_Switch.Dual_Chanel_Monitor.IS := 1, [4].I_Sector_Disable_Switch.Status := 1, [4].O_Unlock_Valve_Left.FeedBack_Type := 1, [4].O_Unlock_Valve_Left.Discrepancy_Time := 3000, [4].O_Unlock_Valve_Left.I_FeedBack_Data := 1, [4].O_Unlock_Valve_Left.I_FeedBack_Status := 1, [4].O_Unlock_Valve_Left.I_Output_Status := 1, [4].O_Unlock_Valve_Right.FeedBack_Type := 1, [4].O_Unlock_Valve_Right.Discrepancy_Time := 3000, [4].O_Unlock_Valve_Right.I_FeedBack_Data := 1, [4].O_Unlock_Valve_Right.I_FeedBack_Status := 1, [4].O_Unlock_Valve_Right.I_Output_Status := 1, [5].Sensors_ChA := 1, [5].Sensors_ChB := 1, [5].LapBar_Open_Close := 1, [5].Input_Status := 1, [5].Sensor_ChA_Open_Memory := 1, [5].Sensor_ChB_Open_Memory := 1, [5].I_LB_PressureSwitch_Valve_Right_Open := 1, [5].I_LB_PressureSwitch_Valve_Left_Open := 1, [5].All_Rack_Memory_Signal_ON := 1, [5].RESTRAINTS_Rack_Sector_ON := 1, [5].I_Close_Position.ChannelA := 1, [5].I_Close_Position.ChannelB := 1, [5].I_Close_Position.InputStatus := 1, [5].I_Close_Position.SafetyFunction := 41, [5].I_Close_Position.DiscrepancyTime := 3000, [5].I_Close_Position.O1 := 1, [5].I_Close_Position.IS := 1, [5].I_Sector_Disable_Switch.Dual_Chanel_Monitor.ChannelB := 1, [5].I_Sector_Disable_Switch.Dual_Chanel_Monitor.InputStatus := 1, [5].I_Sector_Disable_Switch.Dual_Chanel_Monitor.SafetyFunction := 41, [5].I_Sector_Disable_Switch.Dual_Chanel_Monitor.InputType := 2, [5].I_Sector_Disable_Switch.Dual_Chanel_Monitor.DiscrepancyTime := 3000, [5].I_Sector_Disable_Switch.Dual_Chanel_Monitor.IS := 1, [5].I_Sector_Disable_Switch.Status := 1, [5].O_Unlock_Valve_Left.FeedBack_Type := 1, [5].O_Unlock_Valve_Left.Discrepancy_Time := 3000, [5].O_Unlock_Valve_Left.I_FeedBack_Data := 1, [5].O_Unlock_Valve_Left.I_FeedBack_Status := 1, [5].O_Unlock_Valve_Left.I_Output_Status := 1, [5].O_Unlock_Valve_Right.FeedBack_Type := 1, [5].O_Unlock_Valve_Right.Discrepancy_Time := 3000, [5].O_Unlock_Valve_Right.I_FeedBack_Data := 1, [5].O_Unlock_Valve_Right.I_FeedBack_Status := 1, [5].O_Unlock_Valve_Right.I_Output_Status := 1, [6].Sensors_ChA := 1, [6].Sensors_ChB := 1, [6].LapBar_Open_Close := 1, [6].Input_Status := 1, [6].Sensor_ChA_Open_Memory := 1, [6].Sensor_ChB_Open_Memory := 1, [6].I_LB_PressureSwitch_Valve_Right_Open := 1, [6].I_LB_PressureSwitch_Valve_Left_Open := 1, [6].All_Rack_Memory_Signal_ON := 1, [6].RESTRAINTS_Rack_Sector_ON := 1,
